      Appearance <- "SDC\_EDIT"
      ProcessValue <- "DB_SDC_GLOBAL_SYNCH[7].MIN_FAKT"
      ObjectEnable <- "SDC\_EDIT"
   IOField "EA-Feld_95" at 217,452 size 96x29; Authorization "Benutzerverwaltung"; FormatPattern 99999999
      Appearance <- "SDC\_EDIT"
      ProcessValue <- "DB_SDC_GLOBAL_SYNCH[8].HYST"
      ObjectEnable <- "SDC\_EDIT"
   IOField "EA-Feld_96" at 320,452 size 64x29; Authorization "Benutzerverwaltung"; FormatPattern 99.9
      Appearance <- "SDC\_EDIT"
      ProcessValue <- "DB_SDC_GLOBAL_SYNCH[8].K"
      ObjectEnable <- "SDC\_EDIT"
   IOField "EA-Feld_97" at 390,452 size 64x29; Authorization "Benutzerverwaltung"; FormatPattern 99.99
      Appearance <- "SDC\_EDIT"
      ProcessValue <- "DB_SDC_GLOBAL_SYNCH[8].MAX_FAKT"
      ObjectEnable <- "SDC\_EDIT"
   IOField "EA-Feld_98" at 529,452 size 120x29; Authorization "Benutzerverwaltung"; FormatPattern 99999999
      Appearance <- "SDC\_EDIT"
      ProcessValue <- "DB_SDC_GLOBAL_SYNCH[8].SET_DIST"
      ObjectEnable <- "SDC\_EDIT"
   IOField "EA-Feld_99" at 655,452 size 120x29; Authorization "Benutzerverwaltung"; FormatPattern 99999999
      Appearance <- "SDC\_EDIT"
      ProcessValue <- "DB_SDC_GLOBAL_SYNCH[8].SYNCH_DIST"
      ObjectEnable <- "SDC\_EDIT"
   IOField "EA-Feld_100" at 459,452 size 64x29; Authorization "Benutzerverwaltung"; FormatPattern 99.9
      Appearance <- "SDC\_EDIT"
      ProcessValue <- "DB_SDC_GLOBAL_SYNCH[8].MIN_FAKT"
      ObjectEnable <- "SDC\_EDIT"
   IOField "EA-Feld_101" at 217,486 size 96x29; Authorization "Benutzerverwaltung"; FormatPattern 99999999
      Appearance <- "SDC\_EDIT"
      ProcessValue <- "DB_SDC_GLOBAL_SYNCH[9].HYST"
      ObjectEnable <- "SDC\_EDIT"
   IOField "EA-Feld_102" at 320,486 size 64x29; Authorization "Benutzerverwaltung"; FormatPattern 99.9
      Appearance <- "SDC\_EDIT"
      ProcessValue <- "DB_SDC_GLOBAL_SYNCH[9].K"
      ObjectEnable <- "SDC\_EDIT"
   IOField "EA-Feld_103" at 390,486 size 64x29; Authorization "Benutzerverwaltung"; FormatPattern 99.99
      Appearance <- "SDC\_EDIT"
      ProcessValue <- "DB_SDC_GLOBAL_SYNCH[9].MAX_FAKT"
      ObjectEnable <- "SDC\_EDIT"
   IOField "EA-Feld_104" at 529,486 size 120x29; Authorization "Benutzerverwaltung"; FormatPattern 99999999
      Appearance <- "SDC\_EDIT"
      ProcessValue <- "DB_SDC_GLOBAL_SYNCH[9].SET_DIST"
      ObjectEnable <- "SDC\_EDIT"
   IOField "EA-Feld_105" at 655,486 size 120x29; Authorization "Benutzerverwaltung"; FormatPattern 99999999
      Appearance <- "SDC\_EDIT"
      ProcessValue <- "DB_SDC_GLOBAL_SYNCH[9].SYNCH_DIST"
      ObjectEnable <- "SDC\_EDIT"
   IOField "EA-Feld_106" at 459,486 size 64x29; Authorization "Benutzerverwaltung"; FormatPattern 99.9
      Appearance <- "SDC\_EDIT"
      ProcessValue <- "DB_SDC_GLOBAL_SYNCH[9].MIN_FAKT"
      ObjectEnable <- "SDC\_EDIT"
   IOField "EA-Feld_107" at 217,519 size 96x29; Authorization "Benutzerverwaltung"; FormatPattern 99999999
      Appearance <- "SDC\_EDIT"
      ProcessValue <- "DB_SDC_GLOBAL_SYNCH[10].HYST"
      ObjectEnable <- "SDC\_EDIT"
   IOField "EA-Feld_108" at 320,519 size 64x29; Authorization "Benutzerverwaltung"; FormatPattern 99.9
      Appearance <- "SDC\_EDIT"
      ProcessValue <- "DB_SDC_GLOBAL_SYNCH[10].K"
      ObjectEnable <- "SDC\_EDIT"
   IOField "EA-Feld_109" at 390,519 size 64x29; Authorization "Benutzerverwaltung"; FormatPattern 99.99
      Appearance <- "SDC\_EDIT"
      ProcessValue <- "DB_SDC_GLOBAL_SYNCH[10].MAX_FAKT"
      ObjectEnable <- "SDC\_EDIT"
   IOField "EA-Feld_110" at 529,519 size 120x29; Authorization "Benutzerverwaltung"; FormatPattern 99999999
      Appearance <- "SDC\_EDIT"
      ProcessValue <- "DB_SDC_GLOBAL_SYNCH[10].SET_DIST"
      ObjectEnable <- "SDC\_EDIT"
   IOField "EA-Feld_111" at 655,519 size 120x29; Authorization "Benutzerverwaltung"; FormatPattern 99999999
      Appearance <- "SDC\_EDIT"
      ProcessValue <- "DB_SDC_GLOBAL_SYNCH[10].SYNCH_DIST"
      ObjectEnable <- "SDC\_EDIT"
   IOField "EA-Feld_112" at 459,519 size 64x29; Authorization "Benutzerverwaltung"; FormatPattern 99.9
      Appearance <- "SDC\_EDIT"
      ProcessValue <- "DB_SDC_GLOBAL_SYNCH[10].MIN_FAKT"
      ObjectEnable <- "SDC\_EDIT"
   IOField "EA-Feld_113" at 217,553 size 96x29; Authorization "Benutzerverwaltung"; FormatPattern 99999999
      Appearance <- "SDC\_EDIT"
      ProcessValue <- "DB_SDC_GLOBAL_SYNCH[11].HYST"
      ObjectEnable <- "SDC\_EDIT"
   IOField "EA-Feld_114" at 320,553 size 64x29; Authorization "Benutzerverwaltung"; FormatPattern 99.9
      Appearance <- "SDC\_EDIT"
      ProcessValue <- "DB_SDC_GLOBAL_SYNCH[11].K"
      ObjectEnable <- "SDC\_EDIT"
   IOField "EA-Feld_115" at 390,553 size 64x29; Authorization "Benutzerverwaltung"; FormatPattern 99.99
      Appearance <- "SDC\_EDIT"
      ProcessValue <- "DB_SDC_GLOBAL_SYNCH[11].MAX_FAKT"
      ObjectEnable <- "SDC\_EDIT"
   IOField "EA-Feld_116" at 529,553 size 120x29; Authorization "Benutzerverwaltung"; FormatPattern 99999999
      Appearance <- "SDC\_EDIT"
      ProcessValue <- "DB_SDC_GLOBAL_SYNCH[11].SET_DIST"
      ObjectEnable <- "SDC\_EDIT"
   IOField "EA-Feld_117" at 655,553 size 120x29; Authorization "Benutzerverwaltung"; FormatPattern 99999999
      Appearance <- "SDC\_EDIT"
      ProcessValue <- "DB_SDC_GLOBAL_SYNCH[11].SYNCH_DIST"
      ObjectEnable <- "SDC\_EDIT"
   IOField "EA-Feld_118" at 459,553 size 64x29; Authorization "Benutzerverwaltung"; FormatPattern 99.9
      Appearance <- "SDC\_EDIT"
      ProcessValue <- "DB_SDC_GLOBAL_SYNCH[11].MIN_FAKT"
      ObjectEnable <- "SDC\_EDIT"
   IOField "EA-Feld_119" at 217,587 size 96x29; Authorization "Benutzerverwaltung"; FormatPattern 99999999
      Appearance <- "SDC\_EDIT"
      ProcessValue <- "DB_SDC_GLOBAL_SYNCH[12].HYST"
      ObjectEnable <- "SDC\_EDIT"
   IOField "EA-Feld_120" at 320,587 size 64x29; Authorization "Benutzerverwaltung"; FormatPattern 99.9
      Appearance <- "SDC\_EDIT"
      ProcessValue <- "DB_SDC_GLOBAL_SYNCH[12].K"
      ObjectEnable <- "SDC\_EDIT"
   IOField "EA-Feld_121" at 390,587 size 64x29; Authorization "Benutzerverwaltung"; FormatPattern 99.99
      Appearance <- "SDC\_EDIT"
      ProcessValue <- "DB_SDC_GLOBAL_SYNCH[12].MAX_FAKT"
      ObjectEnable <- "SDC\_EDIT"
   IOField "EA-Feld_122" at 529,587 size 120x29; Authorization "Benutzerverwaltung"; FormatPattern 99999999
      Appearance <- "SDC\_EDIT"
      ProcessValue <- "DB_SDC_GLOBAL_SYNCH[12].SET_DIST"
      ObjectEnable <- "SDC\_EDIT"
   IOField "EA-Feld_123" at 655,587 size 120x29; Authorization "Benutzerverwaltung"; FormatPattern 99999999
      Appearance <- "SDC\_EDIT"
      ProcessValue <- "DB_SDC_GLOBAL_SYNCH[12].SYNCH_DIST"
      ObjectEnable <- "SDC\_EDIT"
   IOField "EA-Feld_124" at 459,587 size 64x29; Authorization "Benutzerverwaltung"; FormatPattern 99.9
      Appearance <- "SDC\_EDIT"
      ProcessValue <- "DB_SDC_GLOBAL_SYNCH[12].MIN_FAKT"
      ObjectEnable <- "SDC\_EDIT"
   IOField "EA-Feld_125" at 217,620 size 96x29; Authorization "Benutzerverwaltung"; FormatPattern 99999999
      Appearance <- "SDC\_EDIT"
      ProcessValue <- "DB_SDC_GLOBAL_SYNCH[13].HYST"
      ObjectEnable <- "SDC\_EDIT"
   IOField "EA-Feld_126" at 320,620 size 64x29; Authorization "Benutzerverwaltung"; FormatPattern 99.9
      Appearance <- "SDC\_EDIT"
      ProcessValue <- "DB_SDC_GLOBAL_SYNCH[13].K"
      ObjectEnable <- "SDC\_EDIT"
   IOField "EA-Feld_127" at 390,620 size 64x29; Authorization "Benutzerverwaltung"; FormatPattern 99.99
      Appearance <- "SDC\_EDIT"
      ProcessValue <- "DB_SDC_GLOBAL_SYNCH[13].MAX_FAKT"
      ObjectEnable <- "SDC\_EDIT"
   IOField "EA-Feld_128" at 529,620 size 120x29; Authorization "Benutzerverwaltung"; FormatPattern 99999999
      Appearance <- "SDC\_EDIT"
      ProcessValue <- "DB_SDC_GLOBAL_SYNCH[13].SET_DIST"
      ObjectEnable <- "SDC\_EDIT"
   IOField "EA-Feld_129" at 655,620 size 120x29; Authorization "Benutzerverwaltung"; FormatPattern 99999999
      Appearance <- "SDC\_EDIT"
      ProcessValue <- "DB_SDC_GLOBAL_SYNCH[13].SYNCH_DIST"
      ObjectEnable <- "SDC\_EDIT"
   IOField "EA-Feld_130" at 459,620 size 64x29; Authorization "Benutzerverwaltung"; FormatPattern 99.9
      Appearance <- "SDC\_EDIT"
      ProcessValue <- "DB_SDC_GLOBAL_SYNCH[13].MIN_FAKT"
      ObjectEnable <- "SDC\_EDIT"
   IOField "EA-Feld_131" at 217,654 size 96x29; Authorization "Benutzerverwaltung"; FormatPattern 99999999
      Appearance <- "SDC\_EDIT"
      ProcessValue <- "DB_SDC_GLOBAL_SYNCH[14].HYST"
      ObjectEnable <- "SDC\_EDIT"
   IOField "EA-Feld_132" at 320,654 size 64x29; Authorization "Benutzerverwaltung"; FormatPattern 99.9
      Appearance <- "SDC\_EDIT"
      ProcessValue <- "DB_SDC_GLOBAL_SYNCH[14].K"
      ObjectEnable <- "SDC\_EDIT"
   IOField "EA-Feld_133" at 390,654 size 64x29; Authorization "Benutzerverwaltung"; FormatPattern 99.99
      Appearance <- "SDC\_EDIT"
      ProcessValue <- "DB_SDC_GLOBAL_SYNCH[14].MAX_FAKT"
      ObjectEnable <- "SDC\_EDIT"
   IOField "EA-Feld_134" at 529,654 size 120x29; Authorization "Benutzerverwaltung"; FormatPattern 99999999
      Appearance <- "SDC\_EDIT"
      ProcessValue <- "DB_SDC_GLOBAL_SYNCH[14].SET_DIST"
      ObjectEnable <- "SDC\_EDIT"
   IOField "EA-Feld_135" at 655,654 size 120x29; Authorization "Benutzerverwaltung"; FormatPattern 99999999
      Appearance <- "SDC\_EDIT"
      ProcessValue <- "DB_SDC_GLOBAL_SYNCH[14].SYNCH_DIST"
      ObjectEnable <- "SDC\_EDIT"
   IOField "EA-Feld_136" at 459,654 size 64x29; Authorization "Benutzerverwaltung"; FormatPattern 99.9
      Appearance <- "SDC\_EDIT"
      ProcessValue <- "DB_SDC_GLOBAL_SYNCH[14].MIN_FAKT"
      ObjectEnable <- "SDC\_EDIT"
   IOField "EA-Feld_137" at 217,690 size 96x29; Authorization "Benutzerverwaltung"; FormatPattern 99999999
      Appearance <- "SDC\_EDIT"
      ProcessValue <- "DB_SDC_GLOBAL_SYNCH[15].HYST"
      ObjectEnable <- "SDC\_EDIT"
   IOField "EA-Feld_138" at 320,690 size 64x29; Authorization "Benutzerverwaltung"; FormatPattern 99.9
      Appearance <- "SDC\_EDIT"
      ProcessValue <- "DB_SDC_GLOBAL_SYNCH[15].K"
      ObjectEnable <- "SDC\_EDIT"
   IOField "EA-Feld_139" at 390,690 size 64x29; Authorization "Benutzerverwaltung"; FormatPattern 99.99
      Appearance <- "SDC\_EDIT"
      ProcessValue <- "DB_SDC_GLOBAL_SYNCH[15].MAX_FAKT"
      ObjectEnable <- "SDC\_EDIT"
   IOField "EA-Feld_140" at 529,690 size 120x29; Authorization "Benutzerverwaltung"; FormatPattern 99999999
      Appearance <- "SDC\_EDIT"
      ProcessValue <- "DB_SDC_GLOBAL_SYNCH[15].SET_DIST"
      ObjectEnable <- "SDC\_EDIT"
   IOField "EA-Feld_141" at 655,690 size 120x29; Authorization "Benutzerverwaltung"; FormatPattern 99999999
      Appearance <- "SDC\_EDIT"
      ProcessValue <- "DB_SDC_GLOBAL_SYNCH[15].SYNCH_DIST"
      ObjectEnable <- "SDC\_EDIT"
   IOField "EA-Feld_142" at 459,690 size 64x29; Authorization "Benutzerverwaltung"; FormatPattern 99.9
      Appearance <- "SDC\_EDIT"
      ProcessValue <- "DB_SDC_GLOBAL_SYNCH[15].MIN_FAKT"
      ObjectEnable <- "SDC\_EDIT"
   IOField "EA-Feld_3" at 926,176 size 200x29; Authorization "Benutzerverwaltung"; FormatPattern ????????????????
      Appearance <- "SDC\_EDIT"
      ProcessValue <- "DB_SDC_GLOBAL_REFERENCE_PAR_SET[0].SYNCH"
      ObjectEnable <- "SDC\_EDIT"
   IOField "EA-Feld_4" at 926,210 size 200x29; Authorization "Benutzerverwaltung"; FormatPattern ????????????????
      Appearance <- "SDC\_EDIT"
      ProcessValue <- "DB_SDC_GLOBAL_REFERENCE_PAR_SET[1].SYNCH"
      ObjectEnable <- "SDC\_EDIT"
   IOField "EA-Feld_5" at 926,245 size 200x29; Authorization "Benutzerverwaltung"; FormatPattern ????????????????
      Appearance <- "SDC\_EDIT"
      ProcessValue <- "DB_SDC_GLOBAL_REFERENCE_PAR_SET[2].SYNCH"
      ObjectEnable <- "SDC\_EDIT"
   IOField "EA-Feld_7" at 926,280 size 200x29; Authorization "Benutzerverwaltung"; FormatPattern ????????????????
      Appearance <- "SDC\_EDIT"
      ProcessValue <- "DB_SDC_GLOBAL_REFERENCE_PAR_SET[3].SYNCH"
      ObjectEnable <- "SDC\_EDIT"
   IOField "EA-Feld_8" at 926,314 size 200x29; Authorization "Benutzerverwaltung"; FormatPattern ????????????????
      Appearance <- "SDC\_EDIT"
      ProcessValue <- "DB_SDC_GLOBAL_REFERENCE_PAR_SET[4].SYNCH"
      ObjectEnable <- "SDC\_EDIT"
   IOField "EA-Feld_9" at 926,349 size 200x29; Authorization "Benutzerverwaltung"; FormatPattern ????????????????
      Appearance <- "SDC\_EDIT"
      ProcessValue <- "DB_SDC_GLOBAL_REFERENCE_PAR_SET[5].SYNCH"
      ObjectEnable <- "SDC\_EDIT"
   IOField "EA-Feld_11" at 926,384 size 200x29; Authorization "Benutzerverwaltung"; FormatPattern ????????????????
      Appearance <- "SDC\_EDIT"
      ProcessValue <- "DB_SDC_GLOBAL_REFERENCE_PAR_SET[6].SYNCH"
      ObjectEnable <- "SDC\_EDIT"
   IOField "EA-Feld_13" at 926,418 size 200x29; Authorization "Benutzerverwaltung"; FormatPattern ????????????????
      Appearance <- "SDC\_EDIT"
      ProcessValue <- "DB_SDC_GLOBAL_REFERENCE_PAR_SET[7].SYNCH"
      ObjectEnable <- "SDC\_EDIT"
   IOField "EA-Feld_14" at 926,452 size 200x29; Authorization "Benutzerverwaltung"; FormatPattern ????????????????
      Appearance <- "SDC\_EDIT"
      ProcessValue <- "DB_SDC_GLOBAL_REFERENCE_PAR_SET[8].SYNCH"
      ObjectEnable <- "SDC\_EDIT"
   IOField "EA-Feld_15" at 926,486 size 200x29; Authorization "Benutzerverwaltung"; FormatPattern ????????????????
      Appearance <- "SDC\_EDIT"
      ProcessValue <- "DB_SDC_GLOBAL_REFERENCE_PAR_SET[9].SYNCH"
      ObjectEnable <- "SDC\_EDIT"
   IOField "EA-Feld_16" at 926,519 size 200x29; Authorization "Benutzerverwaltung"; FormatPattern ????????????????
      Appearance <- "SDC\_EDIT"
      ProcessValue <- "DB_SDC_GLOBAL_REFERENCE_PAR_SET[10].SYNCH"
      ObjectEnable <- "SDC\_EDIT"
   IOField "EA-Feld_17" at 926,553 size 200x29; Authorization "Benutzerverwaltung"; FormatPattern ????????????????
      Appearance <- "SDC\_EDIT"
      ProcessValue <- "DB_SDC_GLOBAL_REFERENCE_PAR_SET[11].SYNCH"
      ObjectEnable <- "SDC\_EDIT"
   IOField "EA-Feld_19" at 926,587 size 200x29; Authorization "Benutzerverwaltung"; FormatPattern ????????????????
      Appearance <- "SDC\_EDIT"
      ProcessValue <- "DB_SDC_GLOBAL_REFERENCE_PAR_SET[12].SYNCH"
      ObjectEnable <- "SDC\_EDIT"
   IOField "EA-Feld_20" at 926,620 size 200x29; Authorization "Benutzerverwaltung"; FormatPattern ????????????????
      Appearance <- "SDC\_EDIT"
      ProcessValue <- "DB_SDC_GLOBAL_REFERENCE_PAR_SET[13].SYNCH"
      ObjectEnable <- "SDC\_EDIT"
   IOField "EA-Feld_21" at 926,654 size 200x29; Authorization "Benutzerverwaltung"; FormatPattern ????????????????
      Appearance <- "SDC\_EDIT"
      ProcessValue <- "DB_SDC_GLOBAL_REFERENCE_PAR_SET[14].SYNCH"
      ObjectEnable <- "SDC\_EDIT"
   IOField "EA-Feld_22" at 926,690 size 200x29; Authorization "Benutzerverwaltung"; FormatPattern ????????????????
      Appearance <- "SDC\_EDIT"
      ProcessValue <- "DB_SDC_GLOBAL_REFERENCE_PAR_SET[15].SYNCH"
      ObjectEnable <- "SDC\_EDIT"
   IOField "EA-Feld_143" at 781,176 size 120x30; Authorization "Benutzerverwaltung"; FormatPattern 99999999
      Appearance <- "SDC\_EDIT"
      ProcessValue <- "DB_SDC_GLOBAL_MIN_DIST_EMS[0]"
      ObjectEnable <- "SDC\_EDIT"
   TextField "Textfeld_50" at 769,137 size 119x27; Text 'stop value / Stop Distance / Stop Value'
   IOField "EA-Feld_158" at 781,210 size 120x30; Authorization "Benutzerverwaltung"; FormatPattern 99999999
      Appearance <- "SDC\_EDIT"
      ProcessValue <- "DB_SDC_GLOBAL_MIN_DIST_EMS[1]"
      ObjectEnable <- "SDC\_EDIT"
   IOField "EA-Feld_159" at 781,244 size 120x30; Authorization "Benutzerverwaltung"; FormatPattern 99999999
      Appearance <- "SDC\_EDIT"
      ProcessValue <- "DB_SDC_GLOBAL_MIN_DIST_EMS[2]"
      ObjectEnable <- "SDC\_EDIT"
   IOField "EA-Feld_160" at 781,278 size 120x30; Authorization "Benutzerverwaltung"; FormatPattern 99999999
      Appearance <- "SDC\_EDIT"
      ProcessValue <- "DB_SDC_GLOBAL_MIN_DIST_EMS[3]"
      ObjectEnable <- "SDC\_EDIT"
   IOField "EA-Feld_161" at 781,313 size 120x30; Authorization "Benutzerverwaltung"; FormatPattern 99999999
      Appearance <- "SDC\_EDIT"
      ProcessValue <- "DB_SDC_GLOBAL_MIN_DIST_EMS[4]"
      ObjectEnable <- "SDC\_EDIT"
   IOField "EA-Feld_162" at 781,347 size 120x30; Authorization "Benutzerverwaltung"; FormatPattern 99999999
      Appearance <- "SDC\_EDIT"
      ProcessValue <- "DB_SDC_GLOBAL_MIN_DIST_EMS[5]"
      ObjectEnable <- "SDC\_EDIT"
   IOField "EA-Feld_163" at 781,381 size 120x30; Authorization "Benutzerverwaltung"; FormatPattern 99999999
      Appearance <- "SDC\_EDIT"
      ProcessValue <- "DB_SDC_GLOBAL_MIN_DIST_EMS[6]"
      ObjectEnable <- "SDC\_EDIT"
   IOField "EA-Feld_164" at 781,415 size 120x30; Authorization "Benutzerverwaltung"; FormatPattern 99999999
      Appearance <- "SDC\_EDIT"
      ProcessValue <- "DB_SDC_GLOBAL_MIN_DIST_EMS[7]"
      ObjectEnable <- "SDC\_EDIT"
   IOField "EA-Feld_165" at 781,450 size 120x30; Authorization "Benutzerverwaltung"; FormatPattern 99999999
      Appearance <- "SDC\_EDIT"
      ProcessValue <- "DB_SDC_GLOBAL_MIN_DIST_EMS[8]"
      ObjectEnable <- "SDC\_EDIT"
   IOField "EA-Feld_166" at 781,484 size 120x30; Authorization "Benutzerverwaltung"; FormatPattern 99999999
      Appearance <- "SDC\_EDIT"
      ProcessValue <- "DB_SDC_GLOBAL_MIN_DIST_EMS[9]"
      ObjectEnable <- "SDC\_EDIT"
   IOField "EA-Feld_167" at 781,518 size 120x30; Authorization "Benutzerverwaltung"; FormatPattern 99999999
      Appearance <- "SDC\_EDIT"
      ProcessValue <- "DB_SDC_GLOBAL_MIN_DIST_EMS[10]"
      ObjectEnable <- "SDC\_EDIT"
   IOField "EA-Feld_168" at 781,552 size 120x30; Authorization "Benutzerverwaltung"; FormatPattern 99999999
      Appearance <- "SDC\_EDIT"
      ProcessValue <- "DB_SDC_GLOBAL_MIN_DIST_EMS[11]"
      ObjectEnable <- "SDC\_EDIT"
   IOField "EA-Feld_169" at 781,587 size 120x30; Authorization "Benutzerverwaltung"; FormatPattern 99999999
      Appearance <- "SDC\_EDIT"
      ProcessValue <- "DB_SDC_GLOBAL_MIN_DIST_EMS[12]"
      ObjectEnable <- "SDC\_EDIT"
   IOField "EA-Feld_170" at 781,621 size 120x30; Authorization "Benutzerverwaltung"; FormatPattern 99999999
      Appearance <- "SDC\_EDIT"
      ProcessValue <- "DB_SDC_GLOBAL_MIN_DIST_EMS[13]"
      ObjectEnable <- "SDC\_EDIT"
   IOField "EA-Feld_171" at 781,655 size 120x30; Authorization "Benutzerverwaltung"; FormatPattern 99999999
      Appearance <- "SDC\_EDIT"
      ProcessValue <- "DB_SDC_GLOBAL_MIN_DIST_EMS[14]"
      ObjectEnable <- "SDC\_EDIT"
   IOField "EA-Feld_172" at 781,690 size 120x30; Authorization "Benutzerverwaltung"; FormatPattern 99999999
      Appearance <- "SDC\_EDIT"
      ProcessValue <- "DB_SDC_GLOBAL_MIN_DIST_EMS[15]"
      ObjectEnable <- "SDC\_EDIT"
   TextField "Textfeld_51" at 973,137 size 97x27; Text 'description / Description'
   Button "Schaltfläche_42" at 5,388 size 127x84; TextOff 'EDIT'
      on Click: SetTag("SDC\_EDIT", 0); InvertBit("SDC\_EDIT_BIT")
      Visibility <- "SDC\_EDIT"
      Appearance <- "SDC\_EDIT"

screen "736_DIST_CONTROL_LIMITS_NOT_USED" 1280x800, template "Top_Header"
   on GenerateScreen: SetTag("SDC\_intern_Bildnummer", 736)
   Button "Schaltfläche_2" at 156,142 size 70x593; TextOff 'Text'
   Button "Schaltfläche_1" at 226,142 size 915x42; TextOff 'Text'
   TextField "Textfeld_5" at 172,191 size 35x23; Text '1'
   Button "Schaltfläche_38" at 0,345 size 127x84; TextOff 'EDIT'
      on Click: SetTag("SDC\_EDIT", 1); InvertBit("SDC\_EDIT_BIT")
      Appearance <- "SDC\_EDIT"
   TextField "Textfeld_10" at 172,225 size 35x23; Text '2'
   TextField "Textfeld_14" at 172,259 size 35x23; Text '3'
   TextField "Textfeld_15" at 172,293 size 35x23; Text '4'
   TextField "Textfeld_16" at 172,327 size 35x23; Text '5'
   TextField "Textfeld_17" at 172,361 size 35x23; Text '6'
   TextField "Textfeld_18" at 172,396 size 35x23; Text '7'
   TextField "Textfeld_19" at 172,430 size 35x23; Text '8'
   TextField "Textfeld_20" at 172,464 size 35x23; Text '9'
   TextField "Textfeld_21" at 172,498 size 35x23; Text '10'
   TextField "Textfeld_22" at 164,150 size 58x27; Text 'ParSet'
   TextField "Textfeld_23" at 172,532 size 35x23; Text '11'
   TextField "Textfeld_24" at 172,567 size 35x23; Text '12'
   TextField "Textfeld_25" at 172,601 size 35x23; Text '13'
   TextField "Textfeld_26" at 172,635 size 35x23; Text '14'
   TextField "Textfeld_27" at 172,669 size 35x23; Text '15'
   TextField "Textfeld_28" at 172,704 size 35x23; Text '16'
   TextField "Textfeld_34" at 232,149 size 179x27; Text 'distance slow / Slow Speed Distance'
   IOField "EA-Feld_51" at 244,190 size 170x30; Authorization "Benutzerverwaltung"; FormatPattern 99999999
      Appearance <- "SDC\_EDIT"
      ProcessValue <- "DB_SDC_GLOBAL_LIMITS[0].RAPID_SLOW"
      ObjectEnable <- "SDC\_EDIT"
   IOField "EA-Feld_52" at 611,190 size 170x30; Authorization "Benutzerverwaltung"; FormatPattern 99999999
      Appearance <- "SDC\_EDIT"
      ProcessValue <- "DB_SDC_GLOBAL_MIN_DIST_EMS[0]"
      ObjectEnable <- "SDC\_EDIT"
   IOField "EA-Feld_12" at 481,190 size 64x30; Authorization "Benutzerverwaltung"; FormatPattern 99.9
      Appearance <- "SDC\_EDIT"
      ProcessValue <- "DB_SDC_GLOBAL_LIMITS[0].SLOW_SPEED_FAKT"
      ObjectEnable <- "SDC\_EDIT"
   TextField "Textfeld_40" at 438,149 size 160x27; Text 'coefficient slow / Faktor SlowSpeed / Slow Speed Factor'
   TextField "Textfeld_49" at 609,149 size 425x27; Text 'stop distance (synchron and non synchron area) / Stop Distance (Synchron and Not Synchron Area) / Stop Distance (Synchron and Non Synchron Area)'
   IOField "EA-Feld_3" at 882,188 size 260x30; Authorization "Benutzerverwaltung"; FormatPattern ????????????????
      Appearance <- "SDC\_EDIT"
      ProcessValue <- "DB_SDC_GLOBAL_REFERENCE_PAR_SET[0].LIMITS"
      ObjectEnable <- "SDC\_EDIT"
   IOField "EA-Feld_4" at 882,222 size 260x30; Authorization "Benutzerverwaltung"; FormatPattern ????????????????
      Appearance <- "SDC\_EDIT"
      ProcessValue <- "DB_SDC_GLOBAL_REFERENCE_PAR_SET[1].LIMITS"
      ObjectEnable <- "SDC\_EDIT"
   IOField "EA-Feld_5" at 882,257 size 260x30; Authorization "Benutzerverwaltung"; FormatPattern ????????????????
      Appearance <- "SDC\_EDIT"
      ProcessValue <- "DB_SDC_GLOBAL_REFERENCE_PAR_SET[2].LIMITS"
      ObjectEnable <- "SDC\_EDIT"
   IOField "EA-Feld_7" at 882,292 size 260x30; Authorization "Benutzerverwaltung"; FormatPattern ????????????????
      Appearance <- "SDC\_EDIT"
      ProcessValue <- "DB_SDC_GLOBAL_REFERENCE_PAR_SET[3].LIMITS"
      ObjectEnable <- "SDC\_EDIT"
   IOField "EA-Feld_8" at 882,326 size 260x30; Authorization "Benutzerverwaltung"; FormatPattern ????????????????
      Appearance <- "SDC\_EDIT"
      ProcessValue <- "DB_SDC_GLOBAL_REFERENCE_PAR_SET[4].LIMITS"
      ObjectEnable <- "SDC\_EDIT"
   IOField "EA-Feld_9" at 882,361 size 260x30; Authorization "Benutzerverwaltung"; FormatPattern ????????????????
      Appearance <- "SDC\_EDIT"
      ProcessValue <- "DB_SDC_GLOBAL_REFERENCE_PAR_SET[5].LIMITS"
      ObjectEnable <- "SDC\_EDIT"
   IOField "EA-Feld_11" at 882,396 size 260x30; Authorization "Benutzerverwaltung"; FormatPattern ????????????????
      Appearance <- "SDC\_EDIT"
      ProcessValue <- "DB_SDC_GLOBAL_REFERENCE_PAR_SET[6].LIMITS"
      ObjectEnable <- "SDC\_EDIT"
   IOField "EA-Feld_13" at 882,430 size 260x30; Authorization "Benutzerverwaltung"; FormatPattern ????????????????
      Appearance <- "SDC\_EDIT"
      ProcessValue <- "DB_SDC_GLOBAL_REFERENCE_PAR_SET[7].LIMITS"
      ObjectEnable <- "SDC\_EDIT"
   IOField "EA-Feld_14" at 882,464 size 260x30; Authorization "Benutzerverwaltung"; FormatPattern ????????????????
      Appearance <- "SDC\_EDIT"
      ProcessValue <- "DB_SDC_GLOBAL_REFERENCE_PAR_SET[8].LIMITS"
      ObjectEnable <- "SDC\_EDIT"
   IOField "EA-Feld_15" at 882,498 size 260x30; Authorization "Benutzerverwaltung"; FormatPattern ????????????????
      Appearance <- "SDC\_EDIT"
      ProcessValue <- "DB_SDC_GLOBAL_REFERENCE_PAR_SET[9].LIMITS"
      ObjectEnable <- "SDC\_EDIT"
   IOField "EA-Feld_16" at 882,531 size 260x30; Authorization "Benutzerverwaltung"; FormatPattern ????????????????
      Appearance <- "SDC\_EDIT"
      ProcessValue <- "DB_SDC_GLOBAL_REFERENCE_PAR_SET[10].LIMITS"
      ObjectEnable <- "SDC\_EDIT"
   IOField "EA-Feld_17" at 882,565 size 260x30; Authorization "Benutzerverwaltung"; FormatPattern ????????????????
      Appearance <- "SDC\_EDIT"
      ProcessValue <- "DB_SDC_GLOBAL_REFERENCE_PAR_SET[11].LIMITS"
      ObjectEnable <- "SDC\_EDIT"
   IOField "EA-Feld_19" at 882,599 size 260x30; Authorization "Benutzerverwaltung"; FormatPattern ????????????????
      Appearance <- "SDC\_EDIT"
      ProcessValue <- "DB_SDC_GLOBAL_REFERENCE_PAR_SET[12].LIMITS"
      ObjectEnable <- "SDC\_EDIT"
   IOField "EA-Feld_20" at 882,632 size 260x30; Authorization "Benutzerverwaltung"; FormatPattern ????????????????
      Appearance <- "SDC\_EDIT"
      ProcessValue <- "DB_SDC_GLOBAL_REFERENCE_PAR_SET[13].LIMITS"
      ObjectEnable <- "SDC\_EDIT"
   IOField "EA-Feld_21" at 882,666 size 260x30; Authorization "Benutzerverwaltung"; FormatPattern ????????????????
      Appearance <- "SDC\_EDIT"
      ProcessValue <- "DB_SDC_GLOBAL_REFERENCE_PAR_SET[14].LIMITS"
      ObjectEnable <- "SDC\_EDIT"
   IOField "EA-Feld_22" at 882,702 size 260x30; Authorization "Benutzerverwaltung"; FormatPattern ????????????????
      Appearance <- "SDC\_EDIT"
      ProcessValue <- "DB_SDC_GLOBAL_REFERENCE_PAR_SET[15].LIMITS"
      ObjectEnable <- "SDC\_EDIT"
   IOField "EA-Feld_143" at 244,224 size 170x30; Authorization "Benutzerverwaltung"; FormatPattern 99999999
      Appearance <- "SDC\_EDIT"
      ProcessValue <- "DB_SDC_GLOBAL_LIMITS[1].RAPID_SLOW"
      ObjectEnable <- "SDC\_EDIT"
   IOField "EA-Feld_144" at 244,258 size 170x30; Authorization "Benutzerverwaltung"; FormatPattern 99999999
      Appearance <- "SDC\_EDIT"
      ProcessValue <- "DB_SDC_GLOBAL_LIMITS[2].RAPID_SLOW"
      ObjectEnable <- "SDC\_EDIT"
   IOField "EA-Feld_145" at 244,292 size 170x30; Authorization "Benutzerverwaltung"; FormatPattern 99999999
      Appearance <- "SDC\_EDIT"
      ProcessValue <- "DB_SDC_GLOBAL_LIMITS[3].RAPID_SLOW"
      ObjectEnable <- "SDC\_EDIT"
   IOField "EA-Feld_146" at 244,326 size 170x30; Authorization "Benutzerverwaltung"; FormatPattern 99999999
      Appearance <- "SDC\_EDIT"
      ProcessValue <- "DB_SDC_GLOBAL_LIMITS[4].RAPID_SLOW"
      ObjectEnable <- "SDC\_EDIT"
   IOField "EA-Feld_147" at 244,360 size 170x30; Authorization "Benutzerverwaltung"; FormatPattern 99999999
      Appearance <- "SDC\_EDIT"
      ProcessValue <- "DB_SDC_GLOBAL_LIMITS[5].RAPID_SLOW"
      ObjectEnable <- "SDC\_EDIT"
   IOField "EA-Feld_148" at 244,395 size 170x30; Authorization "Benutzerverwaltung"; FormatPattern 99999999
      Appearance <- "SDC\_EDIT"
      ProcessValue <- "DB_SDC_GLOBAL_LIMITS[6].RAPID_SLOW"
      ObjectEnable <- "SDC\_EDIT"
   IOField "EA-Feld_149" at 244,429 size 170x30; Authorization "Benutzerverwaltung"; FormatPattern 99999999
      Appearance <- "SDC\_EDIT"
      ProcessValue <- "DB_SDC_GLOBAL_LIMITS[7].RAPID_SLOW"
      ObjectEnable <- "SDC\_EDIT"
   IOField "EA-Feld_150" at 244,463 size 170x30; Authorization "Benutzerverwaltung"; FormatPattern 99999999
      Appearance <- "SDC\_EDIT"
      ProcessValue <- "DB_SDC_GLOBAL_LIMITS[8].RAPID_SLOW"
      ObjectEnable <- "SDC\_EDIT"
   IOField "EA-Feld_151" at 244,497 size 170x30; Authorization "Benutzerverwaltung"; FormatPattern 99999999
      Appearance <- "SDC\_EDIT"
      ProcessValue <- "DB_SDC_GLOBAL_LIMITS[9].RAPID_SLOW"
      ObjectEnable <- "SDC\_EDIT"
   IOField "EA-Feld_152" at 244,531 size 170x30; Authorization "Benutzerverwaltung"; FormatPattern 99999999
      Appearance <- "SDC\_EDIT"
      ProcessValue <- "DB_SDC_GLOBAL_LIMITS[10].RAPID_SLOW"
      ObjectEnable <- "SDC\_EDIT"
   IOField "EA-Feld_153" at 244,566 size 170x30; Authorization "Benutzerverwaltung"; FormatPattern 99999999
      Appearance <- "SDC\_EDIT"
      ProcessValue <- "DB_SDC_GLOBAL_LIMITS[11].RAPID_SLOW"
      ObjectEnable <- "SDC\_EDIT"
   IOField "EA-Feld_154" at 244,600 size 170x30; Authorization "Benutzerverwaltung"; FormatPattern 99999999
      Appearance <- "SDC\_EDIT"
      ProcessValue <- "DB_SDC_GLOBAL_LIMITS[12].RAPID_SLOW"
      ObjectEnable <- "SDC\_EDIT"
   IOField "EA-Feld_155" at 244,634 size 170x30; Authorization "Benutzerverwaltung"; FormatPattern 99999999
      Appearance <- "SDC\_EDIT"
      ProcessValue <- "DB_SDC_GLOBAL_LIMITS[13].RAPID_SLOW"
      ObjectEnable <- "SDC\_EDIT"
   IOField "EA-Feld_156" at 244,668 size 170x30; Authorization "Benutzerverwaltung"; FormatPattern 99999999
      Appearance <- "SDC\_EDIT"
      ProcessValue <- "DB_SDC_GLOBAL_LIMITS[14].RAPID_SLOW"
      ObjectEnable <- "SDC\_EDIT"
   IOField "EA-Feld_157" at 244,703 size 170x30; Authorization "Benutzerverwaltung"; FormatPattern 99999999
      Appearance <- "SDC\_EDIT"
      ProcessValue <- "DB_SDC_GLOBAL_LIMITS[15].RAPID_SLOW"
      ObjectEnable <- "SDC\_EDIT"
   IOField "EA-Feld_23" at 481,224 size 64x30; Authorization "Benutzerverwaltung"; FormatPattern 99.9
      Appearance <- "SDC\_EDIT"
      ProcessValue <- "DB_SDC_GLOBAL_LIMITS[1].SLOW_SPEED_FAKT"
      ObjectEnable <- "SDC\_EDIT"
   IOField "EA-Feld_24" at 481,258 size 64x30; Authorization "Benutzerverwaltung"; FormatPattern 99.9
      Appearance <- "SDC\_EDIT"
      ProcessValue <- "DB_SDC_GLOBAL_LIMITS[2].SLOW_SPEED_FAKT"
      ObjectEnable <- "SDC\_EDIT"
   IOField "EA-Feld_25" at 481,292 size 64x30; Authorization "Benutzerverwaltung"; FormatPattern 99.9
      Appearance <- "SDC\_EDIT"
      ProcessValue <- "DB_SDC_GLOBAL_LIMITS[3].SLOW_SPEED_FAKT"
      ObjectEnable <- "SDC\_EDIT"
   IOField "EA-Feld_26" at 481,326 size 64x30; Authorization "Benutzerverwaltung"; FormatPattern 99.9
      Appearance <- "SDC\_EDIT"
      ProcessValue <- "DB_SDC_GLOBAL_LIMITS[4].SLOW_SPEED_FAKT"
      ObjectEnable <- "SDC\_EDIT"
   IOField "EA-Feld_27" at 481,360 size 64x30; Authorization "Benutzerverwaltung"; FormatPattern 99.9
      Appearance <- "SDC\_EDIT"
      ProcessValue <- "DB_SDC_GLOBAL_LIMITS[5].SLOW_SPEED_FAKT"
      ObjectEnable <- "SDC\_EDIT"
   IOField "EA-Feld_28" at 481,395 size 64x30; Authorization "Benutzerverwaltung"; FormatPattern 99.9
      Appearance <- "SDC\_EDIT"
      ProcessValue <- "DB_SDC_GLOBAL_LIMITS[6].SLOW_SPEED_FAKT"
      ObjectEnable <- "SDC\_EDIT"
   IOField "EA-Feld_29" at 481,429 size 64x30; Authorization "Benutzerverwaltung"; FormatPattern 99.9
      Appearance <- "SDC\_EDIT"
      ProcessValue <- "DB_SDC_GLOBAL_LIMITS[7].SLOW_SPEED_FAKT"
      ObjectEnable <- "SDC\_EDIT"
   IOField "EA-Feld_30" at 481,463 size 64x30; Authorization "Benutzerverwaltung"; FormatPattern 99.9
      Appearance <- "SDC\_EDIT"
      ProcessValue <- "DB_SDC_GLOBAL_LIMITS[8].SLOW_SPEED_FAKT"
      ObjectEnable <- "SDC\_EDIT"
   IOField "EA-Feld_31" at 481,497 size 64x30; Authorization "Benutzerverwaltung"; FormatPattern 99.9
      Appearance <- "SDC\_EDIT"
      ProcessValue <- "DB_SDC_GLOBAL_LIMITS[9].SLOW_SPEED_FAKT"
      ObjectEnable <- "SDC\_EDIT"
   IOField "EA-Feld_32" at 481,531 size 64x30; Authorization "Benutzerverwaltung"; FormatPattern 99.9
      Appearance <- "SDC\_EDIT"
      ProcessValue <- "DB_SDC_GLOBAL_LIMITS[10].SLOW_SPEED_FAKT"
      ObjectEnable <- "SDC\_EDIT"
   IOField "EA-Feld_33" at 481,566 size 64x30; Authorization "Benutzerverwaltung"; FormatPattern 99.9
      Appearance <- "SDC\_EDIT"
      ProcessValue <- "DB_SDC_GLOBAL_LIMITS[11].SLOW_SPEED_FAKT"
      ObjectEnable <- "SDC\_EDIT"
   IOField "EA-Feld_34" at 481,600 size 64x30; Authorization "Benutzerverwaltung"; FormatPattern 99.9
      Appearance <- "SDC\_EDIT"
      ProcessValue <- "DB_SDC_GLOBAL_LIMITS[12].SLOW_SPEED_FAKT"
      ObjectEnable <- "SDC\_EDIT"
   IOField "EA-Feld_35" at 481,634 size 64x30; Authorization "Benutzerverwaltung"; FormatPattern 99.9
      Appearance <- "SDC\_EDIT"
      ProcessValue <- "DB_SDC_GLOBAL_LIMITS[13].SLOW_SPEED_FAKT"
      ObjectEnable <- "SDC\_EDIT"
   IOField "EA-Feld_36" at 481,668 size 64x30; Authorization "Benutzerverwaltung"; FormatPattern 99.9
      Appearance <- "SDC\_EDIT"
      ProcessValue <- "DB_SDC_GLOBAL_LIMITS[14].SLOW_SPEED_FAKT"
      ObjectEnable <- "SDC\_EDIT"
   IOField "EA-Feld_37" at 481,703 size 64x30; Authorization "Benutzerverwaltung"; FormatPattern 99.9
      Appearance <- "SDC\_EDIT"
      ProcessValue <- "DB_SDC_GLOBAL_LIMITS[15].SLOW_SPEED_FAKT"
      ObjectEnable <- "SDC\_EDIT"
   IOField "EA-Feld_158" at 611,224 size 170x30; Authorization "Benutzerverwaltung"; FormatPattern 99999999
      Appearance <- "SDC\_EDIT"
      ProcessValue <- "DB_SDC_GLOBAL_MIN_DIST_EMS[1]"
      ObjectEnable <- "SDC\_EDIT"
   IOField "EA-Feld_159" at 611,258 size 170x30; Authorization "Benutzerverwaltung"; FormatPattern 99999999
      Appearance <- "SDC\_EDIT"
      ProcessValue <- "DB_SDC_GLOBAL_MIN_DIST_EMS[2]"
      ObjectEnable <- "SDC\_EDIT"
   IOField "EA-Feld_160" at 611,292 size 170x30; Authorization "Benutzerverwaltung"; FormatPattern 99999999
      Appearance <- "SDC\_EDIT"
      ProcessValue <- "DB_SDC_GLOBAL_MIN_DIST_EMS[3]"
      ObjectEnable <- "SDC\_EDIT"
   IOField "EA-Feld_161" at 611,326 size 170x30; Authorization "Benutzerverwaltung"; FormatPattern 99999999
      Appearance <- "SDC\_EDIT"
      ProcessValue <- "DB_SDC_GLOBAL_MIN_DIST_EMS[4]"
      ObjectEnable <- "SDC\_EDIT"
   IOField "EA-Feld_162" at 611,360 size 170x30; Authorization "Benutzerverwaltung"; FormatPattern 99999999
      Appearance <- "SDC\_EDIT"
      ProcessValue <- "DB_SDC_GLOBAL_MIN_DIST_EMS[5]"
      ObjectEnable <- "SDC\_EDIT"
   IOField "EA-Feld_163" at 611,395 size 170x30; Authorization "Benutzerverwaltung"; FormatPattern 99999999
      Appearance <- "SDC\_EDIT"
      ProcessValue <- "DB_SDC_GLOBAL_MIN_DIST_EMS[6]"
      ObjectEnable <- "SDC\_EDIT"
   IOField "EA-Feld_164" at 611,429 size 170x30; Authorization "Benutzerverwaltung"; FormatPattern 99999999
      Appearance <- "SDC\_EDIT"
      ProcessValue <- "DB_SDC_GLOBAL_MIN_DIST_EMS[7]"
      ObjectEnable <- "SDC\_EDIT"
   IOField "EA-Feld_165" at 611,463 size 170x30; Authorization "Benutzerverwaltung"; FormatPattern 99999999
      Appearance <- "SDC\_EDIT"
      ProcessValue <- "DB_SDC_GLOBAL_MIN_DIST_EMS[8]"
      ObjectEnable <- "SDC\_EDIT"
   IOField "EA-Feld_166" at 611,497 size 170x30; Authorization "Benutzerverwaltung"; FormatPattern 99999999
      Appearance <- "SDC\_EDIT"
      ProcessValue <- "DB_SDC_GLOBAL_MIN_DIST_EMS[9]"
      ObjectEnable <- "SDC\_EDIT"
   IOField "EA-Feld_167" at 611,531 size 170x30; Authorization "Benutzerverwaltung"; FormatPattern 99999999
      Appearance <- "SDC\_EDIT"
      ProcessValue <- "DB_SDC_GLOBAL_MIN_DIST_EMS[10]"
      ObjectEnable <- "SDC\_EDIT"
   IOField "EA-Feld_168" at 611,566 size 170x30; Authorization "Benutzerverwaltung"; FormatPattern 99999999
      Appearance <- "SDC\_EDIT"
      ProcessValue <- "DB_SDC_GLOBAL_MIN_DIST_EMS[11]"
      ObjectEnable <- "SDC\_EDIT"
   IOField "EA-Feld_169" at 611,600 size 170x30; Authorization "Benutzerverwaltung"; FormatPattern 99999999
      Appearance <- "SDC\_EDIT"
      ProcessValue <- "DB_SDC_GLOBAL_MIN_DIST_EMS[12]"
      ObjectEnable <- "SDC\_EDIT"
   IOField "EA-Feld_170" at 611,634 size 170x30; Authorization "Benutzerverwaltung"; FormatPattern 99999999
      Appearance <- "SDC\_EDIT"
      ProcessValue <- "DB_SDC_GLOBAL_MIN_DIST_EMS[13]"
      ObjectEnable <- "SDC\_EDIT"
   IOField "EA-Feld_171" at 611,668 size 170x30; Authorization "Benutzerverwaltung"; FormatPattern 99999999
      Appearance <- "SDC\_EDIT"
      ProcessValue <- "DB_SDC_GLOBAL_MIN_DIST_EMS[14]"
      ObjectEnable <- "SDC\_EDIT"
   IOField "EA-Feld_172" at 611,703 size 170x30; Authorization "Benutzerverwaltung"; FormatPattern 99999999
      Appearance <- "SDC\_EDIT"
      ProcessValue <- "DB_SDC_GLOBAL_MIN_DIST_EMS[15]"
      ObjectEnable <- "SDC\_EDIT"
   Button "Schaltfläche_42" at 0,345 size 127x84; TextOff 'EDIT'
      on Click: SetTag("SDC\_EDIT", 0); InvertBit("SDC\_EDIT_BIT")
      Visibility <- "SDC\_EDIT"
      Appearance <- "SDC\_EDIT"

screen "750_Profinet_Status_NOT_USED" 1280x800, template "Top_Header"
   TextField "Text field_1" at 35,213 size 132x25; Text 'EMS Carrier 1'
   TextField "Text field_2" at 38,380 size 132x25; Text 'EMS Carrier 2'
   TextField "Text field_3" at 35,545 size 132x25; Text 'EMS Carrier 3'
   TextField "Text field_4" at 32,715 size 132x25; Text 'EMS Carrier 4'
   Rectangle "Rectangle_1" at 191,194 size 150x61
      Appearance <- "Carrier 1 G120 D Status"
   TextField "Text field_5" at 206,209 size 131x25; Text 'G120 D Drive'
   Rectangle "Rectangle_2" at 419,194 size 150x61
      Appearance <- "Carrier 1 PnF Encoder Status"
   TextField "Text field_6" at 433,209 size 128x25; Text 'Pn F Encoder'
   Rectangle "Rectangle_3" at 191,363 size 150x61
      Appearance <- "Carrier 2 G120 D Status"
   TextField "Text field_7" at 206,378 size 131x25; Text 'G120 D Drive'
   Rectangle "Rectangle_4" at 419,363 size 150x61
      Appearance <- "Carrier 2 PnF Encoder Status"
   TextField "Text field_8" at 433,378 size 128x25; Text 'Pn F Encoder'
   Rectangle "Rectangle_5" at 191,532 size 150x61
      Appearance <- "Carrier 3  G120 D Status"
   TextField "Text field_9" at 206,547 size 131x25; Text 'G120 D Drive'
   Rectangle "Rectangle_6" at 419,532 size 150x61
      Appearance <- "Carrier 3  PnF Encoder Status"
   TextField "Text field_10" at 433,547 size 128x25; Text 'Pn F Encoder'
   Rectangle "Rectangle_7" at 191,701 size 150x61
      Appearance <- "Carrier 4 G120 D Status"
   TextField "Text field_11" at 206,716 size 131x25; Text 'G120 D Drive'
   Rectangle "Rectangle_8" at 419,701 size 150x61
      Appearance <- "Carrier 4 PnF Encoder Status"
   TextField "Text field_12" at 433,716 size 128x25; Text 'Pn F Encoder'
   Rectangle "Rectangle_9" at 650,194 size 150x61
      Appearance <- "Carrier 1 HMI Status"
   Rectangle "Rectangle_10" at 650,363 size 150x61
      Appearance <- "Carrier 2  HMI Staus"
   Rectangle "Rectangle_11" at 650,532 size 150x61
      Appearance <- "Carrier 3 HMI Status"
   Rectangle "Rectangle_12" at 650,701 size 150x61
      Appearance <- "Carrier 4 HMI Status"
   TextField "Text field_13" at 662,211 size 128x25; Text 'IRD 400 HMI'
   TextField "Text field_14" at 667,380 size 128x25; Text 'IRD 400 HMI'
   TextField "Text field_15" at 662,545 size 128x25; Text 'IRD 400 HMI'
   TextField "Text field_16" at 662,715 size 128x25; Text 'IRD 400 HMI'
   TextField "Text field_17" at 461,144 size 302x26; Text 'Carrier Wise Profinet Diagnosis'
   Rectangle "Rectangle_13" at 878,194 size 150x61
      Appearance <- "Carrier 1 HMI Status"
   TextField "Text field_18" at 915,211 size 79x25; Text 'WLAN 1'
   Rectangle "Rectangle_14" at 878,362 size 150x61
      Appearance <- "Carrier 1 HMI Status"
   TextField "Text field_19" at 915,379 size 79x25; Text 'WLAN 2'
   Rectangle "Rectangle_15" at 878,530 size 150x61
      Appearance <- "Carrier 1 HMI Status"
   TextField "Text field_20" at 915,547 size 79x25; Text 'WLAN 3'
   Rectangle "Rectangle_16" at 878,698 size 150x61
      Appearance <- "Carrier 1 HMI Status"
   TextField "Text field_21" at 915,715 size 79x25; Text 'WLAN 4'
   IOField "EA-Feld_4" at 65,136 size 56x32; FormatPattern 9999
      on OnFinishInput: "SDC_TS_PARAMETER"(); "SDC_TS_REFERENCE"("SDC\_TS_Nr")
      ProcessValue <- "SDC\_TS_Nr"
   TextField "Textfeld_3" at 164,136 size 212x33; Text 'section no. / Sektionnumber / Carrier No'
   Button "Schaltfläche_1" at 122,136 size 40x32; TextOff '+'
      on Click: function_dd21b452("SDC\_TS_Nr", 1); "SDC_TS_PARAMETER"(); "SDC_TS_REFERENCE"("SDC\_TS_Nr")
   Button "Schaltfläche_3" at 25,136 size 39x32; TextOff '-'
      on Click: function_b9b71300("SDC\_TS_Nr", 1); "SDC_TS_PARAMETER"(); "SDC_TS_REFERENCE"("SDC\_TS_Nr")

screen "751_Topic_001.0_PLC" 1280x800, template "Top_Header"
   on GenerateScreen: SetTag("UserDiag_HmiData_actIOSystem", -1)
   on ClearScreen: SetTag("UserDiag_HmiData_actIOSystem", -2)
   TextField "Text field_1" at 29,138 size 51x32; Text 'PLC'
   ScreenModuleView "typeSlot_1" at 292,253 size 49x139; Guid_{11997190-58737} '01'; ScreenModuleType ""
      Guid_{11997190-58740} <- "[1]"
      Guid_{11997190-58743} <- "[1]"
   ScreenModuleView "typeSlot_2" at 245,253 size 49x139; ScreenModuleType ""
      Guid_{11997190-58740} <- "[0]"
      Guid_{11997190-58743} <- "[0]"
   ScreenModuleView "typeSlot_3" at 340,253 size 49x139; Guid_{11997190-58737} '02'; ScreenModuleType ""
      Guid_{11997190-58740} <- "[2]"
      Guid_{11997190-58743} <- "[2]"
   ScreenModuleView "typeSlot_4" at 387,253 size 49x139; Guid_{11997190-58737} '03'; ScreenModuleType ""
      Guid_{11997190-58740} <- "[3]"
      Guid_{11997190-58743} <- "[3]"
   ScreenModuleView "typeSlot_5" at 435,253 size 49x139; Guid_{11997190-58737} '04'; ScreenModuleType ""
      Guid_{11997190-58740} <- "[4]"
      Guid_{11997190-58743} <- "[4]"
   ScreenModuleView "typeSlot_6" at 482,253 size 49x139; Guid_{11997190-58737} '05'; ScreenModuleType ""
      Guid_{11997190-58740} <- "[5]"
      Guid_{11997190-58743} <- "[5]"
   ScreenModuleView "typeSlot_7" at 530,253 size 49x139; Guid_{11997190-58737} '06'; ScreenModuleType ""
      Guid_{11997190-58740} <- "[6]"
      Guid_{11997190-58743} <- "[6]"
   ScreenModuleView "typeSlot_8" at 577,253 size 49x139; Guid_{11997190-58737} '07'; ScreenModuleType ""
      Guid_{11997190-58740} <- "[7]"
      Guid_{11997190-58743} <- "[7]"
   ScreenModuleView "typeSlot_9" at 625,253 size 49x139; Guid_{11997190-58737} '08'; ScreenModuleType ""
      Guid_{11997190-58740} <- "[8]"
      Guid_{11997190-58743} <- "[8]"
   ScreenModuleView "typeSlot_10" at 672,253 size 49x139; Guid_{11997190-58737} '09'; ScreenModuleType ""
      Guid_{11997190-58740} <- "[9]"
      Guid_{11997190-58743} <- "[9]"
   ScreenModuleView "typeSlot_11" at 720,253 size 49x139; Guid_{11997190-58737} '10'; ScreenModuleType ""
      Guid_{11997190-58740} <- "[10]"
      Guid_{11997190-58743} <- "[10]"
   ScreenModuleView "typeSlot_12" at 767,253 size 49x139; Guid_{11997190-58737} '11'; ScreenModuleType ""
      Guid_{11997190-58740} <- "[11]"
      Guid_{11997190-58743} <- "[11]"
   ScreenModuleView "typeSlot_13" at 815,253 size 49x139; Guid_{11997190-58737} '12'; ScreenModuleType ""
      Guid_{11997190-58740} <- "[12]"
      Guid_{11997190-58743} <- "[12]"
   ScreenModuleView "typeSlot_14" at 862,253 size 49x139; Guid_{11997190-58737} '13'; ScreenModuleType ""
      Guid_{11997190-58740} <- "[13]"
      Guid_{11997190-58743} <- "[13]"
   ScreenModuleView "typeSlot_15" at 910,253 size 49x139; Guid_{11997190-58737} '14'; ScreenModuleType ""
      Guid_{11997190-58740} <- "[14]"
      Guid_{11997190-58743} <- "[14]"
   ScreenModuleView "typeSlot_16" at 958,253 size 49x139; Guid_{11997190-58737} '15'; ScreenModuleType ""
      Guid_{11997190-58740} <- "[15]"
      Guid_{11997190-58743} <- "[15]"
   ScreenModuleView "typeSlot_17" at 245,413 size 49x139; Guid_{11997190-58737} '16'; ScreenModuleType ""
      Guid_{11997190-58740} <- "[16]"
      Guid_{11997190-58743} <- "[16]"
   ScreenModuleView "typeSlot_18" at 293,413 size 49x139; Guid_{11997190-58737} '17'; ScreenModuleType ""
      Guid_{11997190-58740} <- "[17]"
      Guid_{11997190-58743} <- "[17]"
   ScreenModuleView "typeSlot_19" at 340,413 size 49x139; Guid_{11997190-58737} '18'; ScreenModuleType ""
      Guid_{11997190-58740} <- "[18]"
      Guid_{11997190-58743} <- "[18]"
   ScreenModuleView "typeSlot_20" at 388,413 size 49x139; Guid_{11997190-58737} '19'; ScreenModuleType ""
      Guid_{11997190-58740} <- "[19]"
      Guid_{11997190-58743} <- "[19]"
   ScreenModuleView "typeSlot_21" at 436,413 size 49x139; Guid_{11997190-58737} '20'; ScreenModuleType ""
      Guid_{11997190-58740} <- "[20]"
      Guid_{11997190-58743} <- "[20]"
   ScreenModuleView "typeSlot_22" at 483,413 size 49x139; Guid_{11997190-58737} '21'; ScreenModuleType ""
      Guid_{11997190-58740} <- "[21]"
      Guid_{11997190-58743} <- "[21]"
   ScreenModuleView "typeSlot_23" at 530,413 size 49x139; Guid_{11997190-58737} '22'; ScreenModuleType ""
      Guid_{11997190-58740} <- "[22]"
      Guid_{11997190-58743} <- "[22]"
   ScreenModuleView "typeSlot_24" at 578,413 size 49x139; Guid_{11997190-58737} '23'; ScreenModuleType ""
      Guid_{11997190-58740} <- "[23]"
      Guid_{11997190-58743} <- "[23]"
   ScreenModuleView "typeSlot_25" at 625,413 size 49x139; Guid_{11997190-58737} '24'; ScreenModuleType ""
      Guid_{11997190-58740} <- "[24]"
      Guid_{11997190-58743} <- "[24]"
   ScreenModuleView "typeSlot_26" at 673,413 size 49x139; Guid_{11997190-58737} '25'; ScreenModuleType ""
      Guid_{11997190-58740} <- "[25]"
      Guid_{11997190-58743} <- "[25]"
   ScreenModuleView "typeSlot_27" at 720,413 size 49x139; Guid_{11997190-58737} '26'; ScreenModuleType ""
      Guid_{11997190-58740} <- "[26]"
      Guid_{11997190-58743} <- "[26]"
   ScreenModuleView "typeSlot_28" at 768,413 size 49x139; Guid_{11997190-58737} '27'; ScreenModuleType ""
      Guid_{11997190-58740} <- "[27]"
      Guid_{11997190-58743} <- "[27]"
   ScreenModuleView "typeSlot_29" at 815,413 size 49x139; Guid_{11997190-58737} '28'; ScreenModuleType ""
      Guid_{11997190-58740} <- "[28]"
      Guid_{11997190-58743} <- "[28]"
   ScreenModuleView "typeSlot_30" at 863,413 size 49x139; Guid_{11997190-58737} '29'; ScreenModuleType ""
      Guid_{11997190-58740} <- "[29]"
      Guid_{11997190-58743} <- "[29]"
   ScreenModuleView "typeSlot_31" at 911,413 size 49x139; Guid_{11997190-58737} '30'; ScreenModuleType ""
      Guid_{11997190-58740} <- "[30]"
      Guid_{11997190-58743} <- "[30]"
   ScreenModuleView "typeSlot_32" at 958,413 size 49x139; Guid_{11997190-58737} '31'; ScreenModuleType ""
      Guid_{11997190-58740} <- "[31]"
      Guid_{11997190-58743} <- "[31]"
   Button "Schaltfläche_64" at 950,700 size 250x80; TextOn 'Reset Übersicht / Reset overview'; TextOff 'Reset Übersicht / Reset overview'
      on Press: function_b14e0dd5("UserDiag_HmiData_ackStates", 0)
   Button "Schaltfläche_3" at 537,578 size 110x80; TextOn 'Legende / Legend'; TextOff 'Legende / Legend'
      on Click: function_efd93a16("Pop-up_Legend", 0, 0, -1, -1, 2)
   IOField "EA-Feld_1" at 550,700 size 80x80; FormatPattern 99; Unit  
      ProcessValue <- "UserDiag_HmiData_ackWaitTime"
   TextField "Textfeld_1" at 260,700 size 277x80; Text 'Wait time Acknowledge [sec] / Wartezeit zur Quittierung'

